      Appearance <- "PN_PB\PTMUX_F_TLN225_240"
   TextField "OBJECT_897" at 258,375 size 40x20; Text '239'
      Appearance <- "PN_PB\PTMUX_F_TLN225_240"
   TextField "OBJECT_905" at 697,420 size 40x20; Text '248'
      Appearance <- "PN_PB\PTMUX_F_TLN241_256"
   TextField "OBJECT_907" at 634,420 size 40x20; Text '249'
      Appearance <- "PN_PB\PTMUX_F_TLN241_256"
   TextField "OBJECT_908" at 571,420 size 40x20; Text '250'
      Appearance <- "PN_PB\PTMUX_F_TLN241_256"
   TextField "OBJECT_909" at 509,420 size 40x20; Text '251'
      Appearance <- "PN_PB\PTMUX_F_TLN241_256"
   TextField "OBJECT_910" at 446,420 size 40x20; Text '252'
      Appearance <- "PN_PB\PTMUX_F_TLN241_256"
   TextField "OBJECT_911" at 383,420 size 40x20; Text '253'
      Appearance <- "PN_PB\PTMUX_F_TLN241_256"
   TextField "OBJECT_912" at 321,420 size 40x20; Text '254'
      Appearance <- "PN_PB\PTMUX_F_TLN241_256"
   TextField "OBJECT_914" at 258,420 size 40x20; Text '255'
      Appearance <- "PN_PB\PTMUX_F_TLN241_256"
   TextField "OBJECT_915" at 885,99 size 40x20; Text '133'
      Appearance <- "PN_PB\PTMUX_F_TLN129_144"
   Group "Group" at 245,86 size 1000x43
   Group "Group_1" at 245,131 size 1000x43
   Group "Group_2" at 245,177 size 1000x43
   Group "Group_3" at 245,222 size 1000x43
   Group "Group_4" at 245,269 size 1000x43
   Group "Group_5" at 245,315 size 1000x43
   Group "Group_6" at 245,362 size 1000x43
   Group "Group_7" at 245,407 size 1000x43
   Button "OBJECT_1046" at 809,86 size 60x43; TextOff 'Text'
      on Press: SetTag("PN_PB\PN\Teiln_Nr", 134)
   Button "OBJECT_1047" at 872,86 size 60x43; TextOff 'Text'
      on Press: SetTag("PN_PB\PN\Teiln_Nr", 133)
   Button "OBJECT_1048" at 935,86 size 60x43; TextOff 'Text'
      on Press: SetTag("PN_PB\PN\Teiln_Nr", 132)
   Button "OBJECT_1049" at 997,86 size 60x43; TextOff 'Text'
      on Press: SetTag("PN_PB\PN\Teiln_Nr", 131)
   Button "OBJECT_1050" at 1060,86 size 60x43; TextOff 'Text'
      on Press: SetTag("PN_PB\PN\Teiln_Nr", 130)
   Button "OBJECT_1051" at 1123,86 size 60x43; TextOff 'Text'
      on Press: SetTag("PN_PB\PN\Teiln_Nr", 129)
   Button "OBJECT_1052" at 1185,86 size 60x43; TextOff 'Text'
      on Press: SetTag("PN_PB\PN\Teiln_Nr", 128)
   Button "OBJECT_1053" at 747,86 size 60x43; TextOff 'Text'
      on Press: SetTag("PN_PB\PN\Teiln_Nr", 135)
   Button "OBJECT_1054" at 684,86 size 60x43; TextOff 'Text'
      on Press: SetTag("PN_PB\PN\Teiln_Nr", 136)
   Button "OBJECT_1055" at 621,86 size 60x43; TextOff 'Text'
      on Press: SetTag("PN_PB\PN\Teiln_Nr", 137)
   Button "OBJECT_1056" at 559,86 size 60x43; TextOff 'Text'
      on Press: SetTag("PN_PB\PN\Teiln_Nr", 138)
   Button "OBJECT_1057" at 496,86 size 60x43; TextOff 'Text'
      on Press: SetTag("PN_PB\PN\Teiln_Nr", 139)
   Button "OBJECT_1058" at 308,86 size 60x43; TextOff 'Text'
      on Press: SetTag("PN_PB\PN\Teiln_Nr", 142)
   Button "OBJECT_1059" at 371,86 size 60x43; TextOff 'Text'
      on Press: SetTag("PN_PB\PN\Teiln_Nr", 141)
   Button "OBJECT_1060" at 433,86 size 60x43; TextOff 'Text'
      on Press: SetTag("PN_PB\PN\Teiln_Nr", 140)
   Button "OBJECT_1061" at 245,86 size 60x43; TextOff 'Text'
      on Press: SetTag("PN_PB\PN\Teiln_Nr", 143)
   Button "OBJECT_1062" at 809,131 size 60x43; TextOff 'Text'
      on Press: SetTag("PN_PB\PN\Teiln_Nr", 150)
   Button "OBJECT_1063" at 872,131 size 60x43; TextOff 'Text'
      on Press: SetTag("PN_PB\PN\Teiln_Nr", 149)
   Button "OBJECT_1064" at 935,131 size 60x43; TextOff 'Text'
      on Press: SetTag("PN_PB\PN\Teiln_Nr", 148)
   Button "OBJECT_1065" at 997,131 size 60x43; TextOff 'Text'
      on Press: SetTag("PN_PB\PN\Teiln_Nr", 147)
   Button "OBJECT_1066" at 1060,131 size 60x43; TextOff 'Text'
      on Press: SetTag("PN_PB\PN\Teiln_Nr", 146)
   Button "OBJECT_1067" at 1123,131 size 60x43; TextOff 'Text'
      on Press: SetTag("PN_PB\PN\Teiln_Nr", 145)
   Button "OBJECT_1068" at 1185,131 size 60x43; TextOff 'Text'
      on Press: SetTag("PN_PB\PN\Teiln_Nr", 144)
   Button "OBJECT_1069" at 747,131 size 60x43; TextOff 'Text'
      on Press: SetTag("PN_PB\PN\Teiln_Nr", 151)
   Button "OBJECT_1070" at 684,131 size 60x43; TextOff 'Text'
      on Press: SetTag("PN_PB\PN\Teiln_Nr", 152)
   Button "OBJECT_1071" at 621,131 size 60x43; TextOff 'Text'
      on Press: SetTag("PN_PB\PN\Teiln_Nr", 153)
   Button "OBJECT_1072" at 559,131 size 60x43; TextOff 'Text'
      on Press: SetTag("PN_PB\PN\Teiln_Nr", 154)
   Button "OBJECT_1073" at 496,131 size 60x43; TextOff 'Text'
      on Press: SetTag("PN_PB\PN\Teiln_Nr", 155)
   Button "OBJECT_1074" at 308,131 size 60x43; TextOff 'Text'
      on Press: SetTag("PN_PB\PN\Teiln_Nr", 158)
   Button "OBJECT_1075" at 371,131 size 60x43; TextOff 'Text'
      on Press: SetTag("PN_PB\PN\Teiln_Nr", 157)
   Button "OBJECT_1076" at 433,131 size 60x43; TextOff 'Text'
      on Press: SetTag("PN_PB\PN\Teiln_Nr", 156)
   Button "OBJECT_1077" at 245,131 size 60x43; TextOff 'Text'
      on Press: SetTag("PN_PB\PN\Teiln_Nr", 159)
   Button "OBJECT_1078" at 809,177 size 60x43; TextOff 'Text'
      on Press: SetTag("PN_PB\PN\Teiln_Nr", 166)
   Button "OBJECT_1079" at 872,177 size 60x43; TextOff 'Text'
      on Press: SetTag("PN_PB\PN\Teiln_Nr", 165)
   Button "OBJECT_1080" at 935,177 size 60x43; TextOff 'Text'
      on Press: SetTag("PN_PB\PN\Teiln_Nr", 164)
   Button "OBJECT_1081" at 997,177 size 60x43; TextOff 'Text'
      on Press: SetTag("PN_PB\PN\Teiln_Nr", 163)
   Button "OBJECT_1082" at 1060,177 size 60x43; TextOff 'Text'
      on Press: SetTag("PN_PB\PN\Teiln_Nr", 162)
   Button "OBJECT_1083" at 1123,177 size 60x43; TextOff 'Text'
      on Press: SetTag("PN_PB\PN\Teiln_Nr", 161)
   Button "OBJECT_1084" at 1185,177 size 60x43; TextOff 'Text'
      on Press: SetTag("PN_PB\PN\Teiln_Nr", 160)
   Button "OBJECT_1085" at 747,177 size 60x43; TextOff 'Text'
      on Press: SetTag("PN_PB\PN\Teiln_Nr", 167)
   Button "OBJECT_1086" at 684,177 size 60x43; TextOff 'Text'
      on Press: SetTag("PN_PB\PN\Teiln_Nr", 168)
   Button "OBJECT_1087" at 621,177 size 60x43; TextOff 'Text'
      on Press: SetTag("PN_PB\PN\Teiln_Nr", 169)
   Button "OBJECT_1088" at 559,177 size 60x43; TextOff 'Text'
      on Press: SetTag("PN_PB\PN\Teiln_Nr", 170)
   Button "OBJECT_1089" at 496,177 size 60x43; TextOff 'Text'
      on Press: SetTag("PN_PB\PN\Teiln_Nr", 171)
   Button "OBJECT_1090" at 308,177 size 60x43; TextOff 'Text'
      on Press: SetTag("PN_PB\PN\Teiln_Nr", 174)
   Button "OBJECT_1091" at 371,177 size 60x43; TextOff 'Text'
      on Press: SetTag("PN_PB\PN\Teiln_Nr", 173)
   Button "OBJECT_1092" at 433,177 size 60x43; TextOff 'Text'
      on Press: SetTag("PN_PB\PN\Teiln_Nr", 172)
   Button "OBJECT_1093" at 245,177 size 60x43; TextOff 'Text'
      on Press: SetTag("PN_PB\PN\Teiln_Nr", 175)
   Button "OBJECT_1094" at 809,222 size 60x43; TextOff 'Text'
      on Press: SetTag("PN_PB\PN\Teiln_Nr", 182)
   Button "OBJECT_1095" at 872,222 size 60x43; TextOff 'Text'
      on Press: SetTag("PN_PB\PN\Teiln_Nr", 181)
   Button "OBJECT_1096" at 935,222 size 60x43; TextOff 'Text'
      on Press: SetTag("PN_PB\PN\Teiln_Nr", 180)
   Button "OBJECT_1097" at 997,222 size 60x43; TextOff 'Text'
      on Press: SetTag("PN_PB\PN\Teiln_Nr", 179)
   Button "OBJECT_1098" at 1060,222 size 60x43; TextOff 'Text'
      on Press: SetTag("PN_PB\PN\Teiln_Nr", 178)
   Button "OBJECT_1099" at 1123,222 size 60x43; TextOff 'Text'
      on Press: SetTag("PN_PB\PN\Teiln_Nr", 177)
   Button "OBJECT_1100" at 1185,222 size 60x43; TextOff 'Text'
      on Press: SetTag("PN_PB\PN\Teiln_Nr", 176)
   Button "OBJECT_1101" at 747,222 size 60x43; TextOff 'Text'
      on Press: SetTag("PN_PB\PN\Teiln_Nr", 183)
   Button "OBJECT_1102" at 684,222 size 60x43; TextOff 'Text'
      on Press: SetTag("PN_PB\PN\Teiln_Nr", 184)
   Button "OBJECT_1103" at 621,222 size 60x43; TextOff 'Text'
      on Press: SetTag("PN_PB\PN\Teiln_Nr", 185)
   Button "OBJECT_1104" at 559,222 size 60x43; TextOff 'Text'
      on Press: SetTag("PN_PB\PN\Teiln_Nr", 186)
   Button "OBJECT_1105" at 496,222 size 60x43; TextOff 'Text'
      on Press: SetTag("PN_PB\PN\Teiln_Nr", 187)
   Button "OBJECT_1106" at 308,222 size 60x43; TextOff 'Text'
      on Press: SetTag("PN_PB\PN\Teiln_Nr", 190)
   Button "OBJECT_1107" at 371,222 size 60x43; TextOff 'Text'
      on Press: SetTag("PN_PB\PN\Teiln_Nr", 189)
   Button "OBJECT_1108" at 433,222 size 60x43; TextOff 'Text'
      on Press: SetTag("PN_PB\PN\Teiln_Nr", 188)
   Button "OBJECT_1109" at 245,222 size 60x43; TextOff 'Text'
      on Press: SetTag("PN_PB\PN\Teiln_Nr", 191)
   Button "OBJECT_1110" at 809,269 size 60x43; TextOff 'Text'
      on Press: SetTag("PN_PB\PN\Teiln_Nr", 198)
   Button "OBJECT_1111" at 872,269 size 60x43; TextOff 'Text'
      on Press: SetTag("PN_PB\PN\Teiln_Nr", 197)
   Button "OBJECT_1112" at 935,269 size 60x43; TextOff 'Text'
      on Press: SetTag("PN_PB\PN\Teiln_Nr", 196)
   Button "OBJECT_1113" at 997,269 size 60x43; TextOff 'Text'
      on Press: SetTag("PN_PB\PN\Teiln_Nr", 195)
   Button "OBJECT_1114" at 1060,269 size 60x43; TextOff 'Text'
      on Press: SetTag("PN_PB\PN\Teiln_Nr", 194)
   Button "OBJECT_1115" at 1123,269 size 60x43; TextOff 'Text'
      on Press: SetTag("PN_PB\PN\Teiln_Nr", 193)
   Button "OBJECT_1116" at 1185,269 size 60x43; TextOff 'Text'
      on Press: SetTag("PN_PB\PN\Teiln_Nr", 192)
   Button "OBJECT_1117" at 747,269 size 60x43; TextOff 'Text'
      on Press: SetTag("PN_PB\PN\Teiln_Nr", 199)
   Button "OBJECT_1118" at 684,269 size 60x43; TextOff 'Text'
      on Press: SetTag("PN_PB\PN\Teiln_Nr", 200)
   Button "OBJECT_1119" at 621,269 size 60x43; TextOff 'Text'
      on Press: SetTag("PN_PB\PN\Teiln_Nr", 201)
   Button "OBJECT_1120" at 559,269 size 60x43; TextOff 'Text'
      on Press: SetTag("PN_PB\PN\Teiln_Nr", 202)
   Button "OBJECT_1121" at 496,269 size 60x43; TextOff 'Text'
      on Press: SetTag("PN_PB\PN\Teiln_Nr", 203)
   Button "OBJECT_1122" at 308,269 size 60x43; TextOff 'Text'
      on Press: SetTag("PN_PB\PN\Teiln_Nr", 206)
   Button "OBJECT_1123" at 371,269 size 60x43; TextOff 'Text'
      on Press: SetTag("PN_PB\PN\Teiln_Nr", 205)
   Button "OBJECT_1124" at 433,269 size 60x43; TextOff 'Text'
      on Press: SetTag("PN_PB\PN\Teiln_Nr", 204)
   Button "OBJECT_1125" at 245,269 size 60x43; TextOff 'Text'
      on Press: SetTag("PN_PB\PN\Teiln_Nr", 207)
   Button "OBJECT_1126" at 809,315 size 60x43; TextOff 'Text'
      on Press: SetTag("PN_PB\PN\Teiln_Nr", 214)
   Button "OBJECT_1127" at 872,315 size 60x43; TextOff 'Text'
      on Press: SetTag("PN_PB\PN\Teiln_Nr", 213)
   Button "OBJECT_1128" at 935,315 size 60x43; TextOff 'Text'
      on Press: SetTag("PN_PB\PN\Teiln_Nr", 212)
   Button "OBJECT_1129" at 997,315 size 60x43; TextOff 'Text'
      on Press: SetTag("PN_PB\PN\Teiln_Nr", 211)
   Button "OBJECT_1130" at 1060,315 size 60x43; TextOff 'Text'
      on Press: SetTag("PN_PB\PN\Teiln_Nr", 210)
   Button "OBJECT_1131" at 1123,315 size 60x43; TextOff 'Text'
      on Press: SetTag("PN_PB\PN\Teiln_Nr", 209)
   Button "OBJECT_1132" at 1185,315 size 60x43; TextOff 'Text'
      on Press: SetTag("PN_PB\PN\Teiln_Nr", 208)
   Button "OBJECT_1133" at 747,315 size 60x43; TextOff 'Text'
      on Press: SetTag("PN_PB\PN\Teiln_Nr", 215)
   Button "OBJECT_1134" at 684,315 size 60x43; TextOff 'Text'
      on Press: SetTag("PN_PB\PN\Teiln_Nr", 216)
   Button "OBJECT_1135" at 621,315 size 60x43; TextOff 'Text'
      on Press: SetTag("PN_PB\PN\Teiln_Nr", 217)
   Button "OBJECT_1136" at 559,315 size 60x43; TextOff 'Text'
      on Press: SetTag("PN_PB\PN\Teiln_Nr", 218)
   Button "OBJECT_1137" at 496,315 size 60x43; TextOff 'Text'
      on Press: SetTag("PN_PB\PN\Teiln_Nr", 219)
   Button "OBJECT_1138" at 308,315 size 60x43; TextOff 'Text'
      on Press: SetTag("PN_PB\PN\Teiln_Nr", 222)
   Button "OBJECT_1139" at 371,315 size 60x43; TextOff 'Text'
      on Press: SetTag("PN_PB\PN\Teiln_Nr", 221)
   Button "OBJECT_1140" at 433,315 size 60x43; TextOff 'Text'
      on Press: SetTag("PN_PB\PN\Teiln_Nr", 220)
   Button "OBJECT_1141" at 245,315 size 60x43; TextOff 'Text'
      on Press: SetTag("PN_PB\PN\Teiln_Nr", 223)
   Button "OBJECT_1142" at 809,362 size 60x43; TextOff 'Text'
      on Press: SetTag("PN_PB\PN\Teiln_Nr", 230)
   Button "OBJECT_1143" at 872,362 size 60x43; TextOff 'Text'
      on Press: SetTag("PN_PB\PN\Teiln_Nr", 229)
   Button "OBJECT_1144" at 935,362 size 60x43; TextOff 'Text'
      on Press: SetTag("PN_PB\PN\Teiln_Nr", 228)
   Button "OBJECT_1145" at 997,362 size 60x43; TextOff 'Text'
      on Press: SetTag("PN_PB\PN\Teiln_Nr", 227)
   Button "OBJECT_1146" at 1060,362 size 60x43; TextOff 'Text'
      on Press: SetTag("PN_PB\PN\Teiln_Nr", 226)
   Button "OBJECT_1147" at 1123,362 size 60x43; TextOff 'Text'
      on Press: SetTag("PN_PB\PN\Teiln_Nr", 225)
   Button "OBJECT_1148" at 1185,362 size 60x43; TextOff 'Text'
      on Press: SetTag("PN_PB\PN\Teiln_Nr", 224)
   Button "OBJECT_1149" at 747,362 size 60x43; TextOff 'Text'
      on Press: SetTag("PN_PB\PN\Teiln_Nr", 231)
   Button "OBJECT_1150" at 684,362 size 60x43; TextOff 'Text'
      on Press: SetTag("PN_PB\PN\Teiln_Nr", 232)
   Button "OBJECT_1151" at 621,362 size 60x43; TextOff 'Text'
      on Press: SetTag("PN_PB\PN\Teiln_Nr", 233)
   Button "OBJECT_1152" at 559,362 size 60x43; TextOff 'Text'
      on Press: SetTag("PN_PB\PN\Teiln_Nr", 234)
   Button "OBJECT_1153" at 496,362 size 60x43; TextOff 'Text'
      on Press: SetTag("PN_PB\PN\Teiln_Nr", 235)
   Button "OBJECT_1154" at 308,362 size 60x43; TextOff 'Text'
      on Press: SetTag("PN_PB\PN\Teiln_Nr", 238)
   Button "OBJECT_1155" at 371,362 size 60x43; TextOff 'Text'
      on Press: SetTag("PN_PB\PN\Teiln_Nr", 237)
   Button "OBJECT_1156" at 433,362 size 60x43; TextOff 'Text'
      on Press: SetTag("PN_PB\PN\Teiln_Nr", 236)
   Button "OBJECT_1157" at 245,362 size 60x43; TextOff 'Text'
      on Press: SetTag("PN_PB\PN\Teiln_Nr", 239)
   Button "OBJECT_1158" at 809,407 size 60x43; TextOff 'Text'
      on Press: SetTag("PN_PB\PN\Teiln_Nr", 246)
   Button "OBJECT_1159" at 872,407 size 60x43; TextOff 'Text'
      on Press: SetTag("PN_PB\PN\Teiln_Nr", 245)
   Button "OBJECT_1160" at 935,407 size 60x43; TextOff 'Text'
      on Press: SetTag("PN_PB\PN\Teiln_Nr", 244)
   Button "OBJECT_1161" at 997,407 size 60x43; TextOff 'Text'
      on Press: SetTag("PN_PB\PN\Teiln_Nr", 243)
   Button "OBJECT_1162" at 1060,407 size 60x43; TextOff 'Text'
      on Press: SetTag("PN_PB\PN\Teiln_Nr", 242)
   Button "OBJECT_1163" at 1123,407 size 60x43; TextOff 'Text'
      on Press: SetTag("PN_PB\PN\Teiln_Nr", 241)
   Button "OBJECT_1164" at 1185,407 size 60x43; TextOff 'Text'
      on Press: SetTag("PN_PB\PN\Teiln_Nr", 240)
   Button "OBJECT_1165" at 747,407 size 60x43; TextOff 'Text'
      on Press: SetTag("PN_PB\PN\Teiln_Nr", 247)
   Button "OBJECT_1166" at 684,407 size 60x43; TextOff 'Text'
      on Press: SetTag("PN_PB\PN\Teiln_Nr", 248)
   Button "OBJECT_1167" at 621,407 size 60x43; TextOff 'Text'
      on Press: SetTag("PN_PB\PN\Teiln_Nr", 249)
   Button "OBJECT_1168" at 559,407 size 60x43; TextOff 'Text'
      on Press: SetTag("PN_PB\PN\Teiln_Nr", 250)
   Button "OBJECT_1169" at 496,407 size 60x43; TextOff 'Text'
      on Press: SetTag("PN_PB\PN\Teiln_Nr", 251)
   Button "OBJECT_1170" at 308,407 size 60x43; TextOff 'Text'
      on Press: SetTag("PN_PB\PN\Teiln_Nr", 254)
   Button "OBJECT_1171" at 371,407 size 60x43; TextOff 'Text'
      on Press: SetTag("PN_PB\PN\Teiln_Nr", 253)
   Button "OBJECT_1172" at 433,407 size 60x43; TextOff 'Text'
      on Press: SetTag("PN_PB\PN\Teiln_Nr", 252)
   Button "OBJECT_1173" at 245,407 size 60x43; TextOff 'Text'
      on Press: SetTag("PN_PB\PN\Teiln_Nr", 255)

screen "100_SDC_PN_Diag0_127" 1280x800, template "SDC"
   on GenerateScreen: SetTag("_intern_BILD_Nr", 100); SetTag("PN_PB\PN\IOSys_ID", 100)
   on ClearScreen: SetTag("_intern_BILD_Nr", 0)
   Button "Schaltfläche_2" at 240,610 size 107x60; TextOff 'Diagnose PN 101'
      on Press: SetTag("PN_PB\PN\IOSys_ID", 101)
      Visibility <- "PN_PB\IO_Sys_ID"
   TextField "OBJECT_21" at 294,46 size 227x27; Text 'ProfiNet-System'
      Visibility <- "PN_PB\IO_Sys_ID"
   TextField "OBJECT_511" at 248,475 size 227x27; Text 'ProfiNet-Teilnehmer:'
      Visibility <- "PN_PB\IO_Sys_ID"
   Button "Schaltfläche_1" at 240,610 size 107x60; TextOff 'Diagnose PN 100'
      on Press: SetTag("PN_PB\PN\IOSys_ID", 100)
      Visibility <- "PN_PB\IO_Sys_ID"
   Button "Schaltfläche_3" at 588,45 size 322x37; TextOff 'ProfiNet-Teilnehmer 128 - 255'
      on Release: ActivateScreen("101_SDC_PN_Diag128_255", 0)
   Button "OBJECT_655" at 1186,89 size 60x40; TextOff 'Text'
      on Press: SetTag("PN_PB\PN\Teiln_Nr", 1)
   GraphicIOField "OBJECT_41" at 936,89 size 60x43; PictureList "PB_Slave_Bit12_2"
      ProcessValue <- "PN_PB\PTMUX_P_TLN1_16"
   GraphicIOField "302" at 309,89 size 60x43; PictureList "PB_Slave_Bit6_2"
      ProcessValue <- "PN_PB\PTMUX_P_TLN1_16"
   GraphicView "OBJECT_496" at 1193,498 size 60x43; Picture "PB_Array_blau_2"
   TextField "OBJECT_497" at 1206,510 size 40x20; Text '1'
   GraphicView "OBJECT_498" at 1193,545 size 60x43; Picture "PB_Array_grün_2"
   TextField "OBJECT_499" at 1206,556 size 40x20; Text '1'
   TextField "OBJECT_500" at 1206,600 size 40x20; Text '1'
   GraphicView "OBJECT_501" at 1193,590 size 60x43; Picture "PB_Array_grün_2"
   TextField "OBJECT_502" at 1206,600 size 40x20; Text '1'
   TextField "OBJECT_504" at 939,505 size 257x31; Text 'Teilnehmer nicht vorhanden'
   TextField "OBJECT_505" at 939,597 size 193x33; Text 'Teilnehmer gestört'
   TextField "OBJECT_506" at 939,552 size 213x33; Text 'Teilnehmer vorhanden'
   GraphicIOField "OBJECT_193" at 748,89 size 60x43; PictureList "PB_Slave_Bit15_2"
      ProcessValue <- "PN_PB\PTMUX_P_TLN1_16"
   GraphicIOField "OBJECT_195" at 810,89 size 60x43; PictureList "PB_Slave_Bit14_2"
      ProcessValue <- "PN_PB\PTMUX_P_TLN1_16"
   TextField "OBJECT_201" at 1009,94 size 40x20; Text '1'
   GraphicIOField "OBJECT_202" at 1061,89 size 60x43; PictureList "PB_Slave_Bit10_2"
      ProcessValue <- "PN_PB\PTMUX_P_TLN1_16"
   GraphicIOField "OBJECT_204" at 1124,89 size 60x43; PictureList "PB_Slave_Bit9_2"
      ProcessValue <- "PN_PB\PTMUX_P_TLN1_16"
   GraphicIOField "OBJECT_205" at 1186,89 size 60x43; PictureList "PB_Slave_Bit8_2"
      ProcessValue <- "PN_PB\PTMUX_P_TLN1_16"
   GraphicIOField "OBJECT_208" at 998,89 size 60x43; PictureList "PB_Slave_Bit11_2"
      ProcessValue <- "PN_PB\PTMUX_P_TLN1_16"
   TextField "OBJECT_233" at 1197,100 size 40x20; Text '0'
      Appearance <- "PN_PB\PTMUX_F_TLN1_16"
   TextField "OBJECT_234" at 1134,100 size 40x20; Text '1'
      Appearance <- "PN_PB\PTMUX_F_TLN1_16"
   TextField "OBJECT_235" at 1072,100 size 40x20; Text '2'
      Appearance <- "PN_PB\PTMUX_F_TLN1_16"
   TextField "OBJECT_236" at 1009,100 size 40x20; Text '3'
      Appearance <- "PN_PB\PTMUX_F_TLN1_16"
   TextField "OBJECT_237" at 946,100 size 40x20; Text '4'
      Appearance <- "PN_PB\PTMUX_F_TLN1_16"
   TextField "OBJECT_239" at 821,100 size 40x20; Text '6'
      Appearance <- "PN_PB\PTMUX_F_TLN1_16"
   TextField "OBJECT_240" at 758,100 size 40x20; Text '7'
      Appearance <- "PN_PB\PTMUX_F_TLN1_16"
   GraphicIOField "OBJECT_241" at 748,134 size 60x43; PictureList "PB_Slave_Bit15_2"
      ProcessValue <- "PN_PB\PTMUX_P_TLN17_32"
   GraphicIOField "OBJECT_242" at 810,134 size 60x43; PictureList "PB_Slave_Bit14_2"
      ProcessValue <- "PN_PB\PTMUX_P_TLN17_32"
   GraphicIOField "OBJECT_243" at 873,134 size 60x43; PictureList "PB_Slave_Bit13_2"
      ProcessValue <- "PN_PB\PTMUX_P_TLN17_32"
   GraphicIOField "OBJECT_244" at 936,134 size 60x43; PictureList "PB_Slave_Bit12_2"
      ProcessValue <- "PN_PB\PTMUX_P_TLN17_32"
   TextField "OBJECT_245" at 1009,145 size 40x20; Text '1'
   GraphicIOField "OBJECT_246" at 1061,134 size 60x43; PictureList "PB_Slave_Bit10_2"
      ProcessValue <- "PN_PB\PTMUX_P_TLN17_32"
   GraphicIOField "OBJECT_247" at 1124,134 size 60x43; PictureList "PB_Slave_Bit9_2"
      ProcessValue <- "PN_PB\PTMUX_P_TLN17_32"
   GraphicIOField "OBJECT_248" at 1186,134 size 60x43; PictureList "PB_Slave_Bit8_2"
      ProcessValue <- "PN_PB\PTMUX_P_TLN17_32"
   GraphicIOField "OBJECT_249" at 998,134 size 60x43; PictureList "PB_Slave_Bit11_2"
      ProcessValue <- "PN_PB\PTMUX_P_TLN17_32"
   TextField "OBJECT_267" at 1134,145 size 40x20; Text '17'
      Appearance <- "PN_PB\PTMUX_F_TLN17_32"
   TextField "OBJECT_268" at 1072,145 size 40x20; Text '18'
      Appearance <- "PN_PB\PTMUX_F_TLN17_32"
   TextField "OBJECT_269" at 1009,145 size 40x20; Text '19'
      Appearance <- "PN_PB\PTMUX_F_TLN17_32"
   TextField "OBJECT_270" at 946,145 size 40x20; Text '20'
      Appearance <- "PN_PB\PTMUX_F_TLN17_32"
   TextField "OBJECT_271" at 884,145 size 40x20; Text '21'
      Appearance <- "PN_PB\PTMUX_F_TLN17_32"
   TextField "OBJECT_272" at 821,145 size 40x20; Text '22'
      Appearance <- "PN_PB\PTMUX_F_TLN17_32"
   TextField "OBJECT_273" at 758,145 size 40x20; Text '23'
      Appearance <- "PN_PB\PTMUX_F_TLN17_32"
   TextField "OBJECT_274" at 1197,145 size 40x20; Text '16'
      Appearance <- "PN_PB\PTMUX_F_TLN17_32"
   GraphicIOField "OBJECT_275" at 748,180 size 60x43; PictureList "PB_Slave_Bit15_2"
      ProcessValue <- "PN_PB\PTMUX_P_TLN33_48"
   GraphicIOField "OBJECT_276" at 873,180 size 60x43; PictureList "PB_Slave_Bit13_2"
      ProcessValue <- "PN_PB\PTMUX_P_TLN33_48"
   GraphicIOField "OBJECT_277" at 936,180 size 60x43; PictureList "PB_Slave_Bit12_2"
      ProcessValue <- "PN_PB\PTMUX_P_TLN33_48"
   TextField "OBJECT_278" at 1009,190 size 40x20; Text '1'
   GraphicIOField "OBJECT_279" at 1061,180 size 60x43; PictureList "PB_Slave_Bit10_2"
      ProcessValue <- "PN_PB\PTMUX_P_TLN33_48"
   GraphicIOField "OBJECT_280" at 1124,180 size 60x43; PictureList "PB_Slave_Bit9_2"
      ProcessValue <- "PN_PB\PTMUX_P_TLN33_48"
   GraphicIOField "OBJECT_281" at 1186,180 size 60x43; PictureList "PB_Slave_Bit8_2"
      ProcessValue <- "PN_PB\PTMUX_P_TLN33_48"
   GraphicIOField "OBJECT_282" at 998,180 size 60x43; PictureList "PB_Slave_Bit11_2"
      ProcessValue <- "PN_PB\PTMUX_P_TLN33_48"
   TextField "OBJECT_300" at 1197,190 size 40x20; Text '32'
      Appearance <- "PN_PB\PTMUX_F_TLN33_48"
   TextField "OBJECT_301" at 1134,190 size 40x20; Text '33'
      Appearance <- "PN_PB\PTMUX_F_TLN33_48"
   TextField "OBJECT_302" at 1072,190 size 40x20; Text '34'
      Appearance <- "PN_PB\PTMUX_F_TLN33_48"
   TextField "OBJECT_303" at 1009,190 size 40x20; Text '35'
      Appearance <- "PN_PB\PTMUX_F_TLN33_48"
   TextField "OBJECT_304" at 946,190 size 40x20; Text '36'
      Appearance <- "PN_PB\PTMUX_F_TLN33_48"
   TextField "OBJECT_305" at 884,190 size 40x20; Text '37'
      Appearance <- "PN_PB\PTMUX_F_TLN33_48"
   TextField "OBJECT_307" at 758,190 size 40x20; Text '39'
      Appearance <- "PN_PB\PTMUX_F_TLN33_48"
   GraphicIOField "OBJECT_308" at 810,180 size 60x43; PictureList "PB_Slave_Bit14_2"
      ProcessValue <- "PN_PB\PTMUX_P_TLN33_48"
   TextField "OBJECT_309" at 821,190 size 40x20; Text '38'
      Appearance <- "PN_PB\PTMUX_F_TLN33_48"
   GraphicIOField "OBJECT_310" at 748,225 size 60x43; PictureList "PB_Slave_Bit15_2"
      ProcessValue <- "PN_PB\PTMUX_P_TLN49_64"
   GraphicIOField "OBJECT_311" at 873,225 size 60x43; PictureList "PB_Slave_Bit13_2"
      ProcessValue <- "PN_PB\PTMUX_P_TLN49_64"
   GraphicIOField "OBJECT_312" at 936,225 size 60x43; PictureList "PB_Slave_Bit12_2"
      ProcessValue <- "PN_PB\PTMUX_P_TLN49_64"
   TextField "OBJECT_313" at 1009,236 size 40x20; Text '1'
   GraphicIOField "OBJECT_314" at 1061,225 size 60x43; PictureList "PB_Slave_Bit10_2"
      ProcessValue <- "PN_PB\PTMUX_P_TLN49_64"
   GraphicIOField "OBJECT_315" at 1124,225 size 60x43; PictureList "PB_Slave_Bit9_2"
      ProcessValue <- "PN_PB\PTMUX_P_TLN49_64"
   GraphicIOField "OBJECT_316" at 1186,225 size 60x43; PictureList "PB_Slave_Bit8_2"
      ProcessValue <- "PN_PB\PTMUX_P_TLN49_64"
   GraphicIOField "OBJECT_317" at 998,225 size 60x43; PictureList "PB_Slave_Bit11_2"
      ProcessValue <- "PN_PB\PTMUX_P_TLN49_64"
   TextField "OBJECT_335" at 1197,236 size 40x20; Text '48'
      Appearance <- "PN_PB\PTMUX_F_TLN49_64"
   TextField "OBJECT_336" at 1134,236 size 40x20; Text '49'
      Appearance <- "PN_PB\PTMUX_F_TLN49_64"
   TextField "OBJECT_337" at 1072,236 size 40x20; Text '50'
      Appearance <- "PN_PB\PTMUX_F_TLN49_64"
   TextField "OBJECT_338" at 946,236 size 40x20; Text '52'
      Appearance <- "PN_PB\PTMUX_F_TLN49_64"
   TextField "OBJECT_339" at 884,236 size 40x20; Text '53'
      Appearance <- "PN_PB\PTMUX_F_TLN49_64"
   TextField "OBJECT_341" at 758,236 size 40x20; Text '55'
      Appearance <- "PN_PB\PTMUX_F_TLN49_64"
   GraphicIOField "OBJECT_342" at 810,225 size 60x43; PictureList "PB_Slave_Bit14_2"
      ProcessValue <- "PN_PB\PTMUX_P_TLN49_64"
   TextField "OBJECT_343" at 821,236 size 40x20; Text '54'
      Appearance <- "PN_PB\PTMUX_F_TLN49_64"
   TextField "OBJECT_344" at 1009,236 size 40x20; Text '51'
      Appearance <- "PN_PB\PTMUX_F_TLN49_64"
   GraphicIOField "OBJECT_345" at 748,270 size 60x43; PictureList "PB_Slave_Bit15_2"
      ProcessValue <- "PN_PB\PTMUX_P_TLN65_80"
   GraphicIOField "OBJECT_346" at 873,270 size 60x43; PictureList "PB_Slave_Bit13_2"
      ProcessValue <- "PN_PB\PTMUX_P_TLN65_80"
   TextField "OBJECT_347" at 1009,282 size 40x20; Text '1'
   GraphicIOField "OBJECT_348" at 1061,270 size 60x43; PictureList "PB_Slave_Bit10_2"
      ProcessValue <- "PN_PB\PTMUX_P_TLN65_80"
   GraphicIOField "OBJECT_349" at 1124,270 size 60x43; PictureList "PB_Slave_Bit9_2"
      ProcessValue <- "PN_PB\PTMUX_P_TLN65_80"
   GraphicIOField "OBJECT_350" at 1186,270 size 60x43; PictureList "PB_Slave_Bit8_2"
      ProcessValue <- "PN_PB\PTMUX_P_TLN65_80"
   GraphicIOField "OBJECT_351" at 998,270 size 60x43; PictureList "PB_Slave_Bit11_2"
      ProcessValue <- "PN_PB\PTMUX_P_TLN65_80"
   TextField "OBJECT_369" at 1197,282 size 40x20; Text '64'
      Appearance <- "PN_PB\PTMUX_F_TLN65_80"
   TextField "OBJECT_370" at 1134,282 size 40x20; Text '65'
      Appearance <- "PN_PB\PTMUX_F_TLN65_80"
   TextField "OBJECT_371" at 1072,282 size 40x20; Text '66'
      Appearance <- "PN_PB\PTMUX_F_TLN65_80"
   TextField "OBJECT_373" at 884,282 size 40x20; Text '69'
      Appearance <- "PN_PB\PTMUX_F_TLN65_80"
   TextField "OBJECT_375" at 758,282 size 40x20; Text '71'
      Appearance <- "PN_PB\PTMUX_F_TLN65_80"
   GraphicIOField "OBJECT_376" at 810,270 size 60x43; PictureList "PB_Slave_Bit14_2"
      ProcessValue <- "PN_PB\PTMUX_P_TLN65_80"
   TextField "OBJECT_377" at 821,282 size 40x20; Text '70'
      Appearance <- "PN_PB\PTMUX_F_TLN65_80"
   TextField "OBJECT_378" at 1009,282 size 40x20; Text '67'
      Appearance <- "PN_PB\PTMUX_F_TLN65_80"
   GraphicIOField "OBJECT_379" at 936,270 size 60x43; PictureList "PB_Slave_Bit12_2"
      ProcessValue <- "PN_PB\PTMUX_P_TLN65_80"
   TextField "OBJECT_380" at 946,282 size 40x20; Text '68'
      Appearance <- "PN_PB\PTMUX_F_TLN65_80"
   GraphicIOField "OBJECT_381" at 748,317 size 60x43; PictureList "PB_Slave_Bit15_2"
      ProcessValue <- "PN_PB\PTMUX_P_TLN81_96"
   GraphicIOField "OBJECT_382" at 873,317 size 60x43; PictureList "PB_Slave_Bit13_2"
      ProcessValue <- "PN_PB\PTMUX_P_TLN81_96"
   TextField "OBJECT_383" at 1009,329 size 40x20; Text '1'
   GraphicIOField "OBJECT_384" at 1061,317 size 60x43; PictureList "PB_Slave_Bit10_2"
      ProcessValue <- "PN_PB\PTMUX_P_TLN81_96"
   GraphicIOField "OBJECT_385" at 1124,317 size 60x43; PictureList "PB_Slave_Bit9_2"
      ProcessValue <- "PN_PB\PTMUX_P_TLN81_96"
   GraphicIOField "OBJECT_386" at 1186,317 size 60x43; PictureList "PB_Slave_Bit8_2"
      ProcessValue <- "PN_PB\PTMUX_P_TLN81_96"
   GraphicIOField "OBJECT_387" at 998,317 size 60x43; PictureList "PB_Slave_Bit11_2"
      ProcessValue <- "PN_PB\PTMUX_P_TLN81_96"
   TextField "OBJECT_405" at 1197,329 size 40x20; Text '80'
      Appearance <- "PN_PB\PTMUX_F_TLN81_96"
   TextField "OBJECT_406" at 1134,329 size 40x20; Text '81'
      Appearance <- "PN_PB\PTMUX_F_TLN81_96"
   TextField "OBJECT_407" at 1072,329 size 40x20; Text '82'
      Appearance <- "PN_PB\PTMUX_F_TLN81_96"
   TextField "OBJECT_409" at 884,329 size 40x20; Text '85'
      Appearance <- "PN_PB\PTMUX_F_TLN81_96"
   GraphicIOField "OBJECT_411" at 810,317 size 60x43; PictureList "PB_Slave_Bit14_2"
      ProcessValue <- "PN_PB\PTMUX_P_TLN81_96"
   TextField "OBJECT_412" at 821,329 size 40x20; Text '86'
      Appearance <- "PN_PB\PTMUX_F_TLN81_96"
   TextField "OBJECT_413" at 1009,329 size 40x20; Text '83'
      Appearance <- "PN_PB\PTMUX_F_TLN81_96"
   GraphicIOField "OBJECT_414" at 936,317 size 60x43; PictureList "PB_Slave_Bit12_2"
      ProcessValue <- "PN_PB\PTMUX_P_TLN81_96"
   TextField "OBJECT_415" at 946,329 size 40x20; Text '84'
      Appearance <- "PN_PB\PTMUX_F_TLN81_96"
   TextField "OBJECT_416" at 758,329 size 40x20; Text '87'
      Appearance <- "PN_PB\PTMUX_F_TLN81_96"
   GraphicIOField "OBJECT_417" at 873,364 size 60x43; PictureList "PB_Slave_Bit13_2"
      ProcessValue <- "PN_PB\PTMUX_P_TLN97_112"
   TextField "OBJECT_418" at 1009,376 size 40x20; Text '1'
   GraphicIOField "OBJECT_419" at 1061,364 size 60x43; PictureList "PB_Slave_Bit10_2"
      ProcessValue <- "PN_PB\PTMUX_P_TLN97_112"
   GraphicIOField "OBJECT_420" at 1124,364 size 60x43; PictureList "PB_Slave_Bit9_2"
      ProcessValue <- "PN_PB\PTMUX_P_TLN97_112"
   GraphicIOField "OBJECT_421" at 1186,364 size 60x43; PictureList "PB_Slave_Bit8_2"
      ProcessValue <- "PN_PB\PTMUX_P_TLN97_112"
   GraphicIOField "OBJECT_422" at 998,364 size 60x43; PictureList "PB_Slave_Bit11_2"
      ProcessValue <- "PN_PB\PTMUX_P_TLN97_112"
   TextField "OBJECT_440" at 1197,376 size 40x20; Text '96'
      Appearance <- "PN_PB\PTMUX_F_TLN97_112"
   TextField "OBJECT_441" at 1134,376 size 40x20; Text '97'
      Appearance <- "PN_PB\PTMUX_F_TLN97_112"
   TextField "OBJECT_442" at 1072,376 size 40x20; Text '98'
      Appearance <- "PN_PB\PTMUX_F_TLN97_112"
   TextField "OBJECT_444" at 884,376 size 40x20; Text '101'
      Appearance <- "PN_PB\PTMUX_F_TLN97_112"
   GraphicIOField "OBJECT_446" at 810,364 size 60x43; PictureList "PB_Slave_Bit14_2"
      ProcessValue <- "PN_PB\PTMUX_P_TLN97_112"
   TextField "OBJECT_447" at 821,376 size 40x20; Text '102'
      Appearance <- "PN_PB\PTMUX_F_TLN97_112"
   TextField "OBJECT_448" at 1009,376 size 40x20; Text '99'
      Appearance <- "PN_PB\PTMUX_F_TLN97_112"
   GraphicIOField "OBJECT_449" at 936,364 size 60x43; PictureList "PB_Slave_Bit12_2"
      ProcessValue <- "PN_PB\PTMUX_P_TLN97_112"
   TextField "OBJECT_450" at 946,376 size 40x20; Text '100'
      Appearance <- "PN_PB\PTMUX_F_TLN97_112"
   GraphicIOField "OBJECT_452" at 748,364 size 60x43; PictureList "PB_Slave_Bit15_2"
      ProcessValue <- "PN_PB\PTMUX_P_TLN97_112"
   TextField "OBJECT_453" at 758,376 size 40x20; Text '103'
      Appearance <- "PN_PB\PTMUX_F_TLN97_112"
   GraphicIOField "OBJECT_454" at 873,410 size 60x43; PictureList "PB_Slave_Bit13_2"
      ProcessValue <- "PN_PB\PTMUX_P_TLN113_128"
   TextField "OBJECT_455" at 1009,421 size 40x20; Text '1'
   GraphicIOField "OBJECT_456" at 1061,410 size 60x43; PictureList "PB_Slave_Bit10_2"
      ProcessValue <- "PN_PB\PTMUX_P_TLN113_128"
   GraphicIOField "OBJECT_457" at 1124,410 size 60x43; PictureList "PB_Slave_Bit9_2"
      ProcessValue <- "PN_PB\PTMUX_P_TLN113_128"
   GraphicIOField "OBJECT_458" at 1186,410 size 60x43; PictureList "PB_Slave_Bit8_2"
      ProcessValue <- "PN_PB\PTMUX_P_TLN113_128"
   GraphicIOField "OBJECT_459" at 998,410 size 60x43; PictureList "PB_Slave_Bit11_2"
      ProcessValue <- "PN_PB\PTMUX_P_TLN113_128"
   TextField "OBJECT_476" at 1197,421 size 40x20; Text '112'
      Appearance <- "PN_PB\PTMUX_F_TLN113_128"
   TextField "OBJECT_477" at 1134,421 size 40x20; Text '113'
      Appearance <- "PN_PB\PTMUX_F_TLN113_128"
   TextField "OBJECT_478" at 1072,421 size 40x20; Text '114'
      Appearance <- "PN_PB\PTMUX_F_TLN113_128"
   TextField "OBJECT_480" at 884,421 size 40x20; Text '117'
      Appearance <- "PN_PB\PTMUX_F_TLN113_128"
   GraphicIOField "OBJECT_482" at 810,410 size 60x43; PictureList "PB_Slave_Bit14_2"
      ProcessValue <- "PN_PB\PTMUX_P_TLN113_128"
   TextField "OBJECT_483" at 821,421 size 40x20; Text '118'